(* Logix 5000 project; controller PLC_MCC1201_220AP1 vendor 1 type 14 code 164 rev 35.11; software revision 35.00 *)

TASK _18_STI (periodic, rate 10 ms, priority 10, watchdog 500 ms) : _18_STI
TASK Diagnostic (periodic, rate 500 ms, priority 15, watchdog 2000 ms) : Modules
TASK MainTask (periodic, rate 10 ms, priority 10, watchdog 500 ms) : MainProgram, CommandLogic

MODULES
   Local : vendor 1 type 14 code 164 (ICP 1, rev 35.11)
      PLC_MCC1300_TEST : vendor 1 type 14 code 166 (Ethernet 192.168.38.1, rev 35.1, $337b92f8$ RPI 20 ms)
      ETH_MCC1201 : 1756-EN2T (ICP 3, Ethernet 138.84.12.111, rev 11.1)
         Cullet_System : vendor 1 type 14 code 164 (Ethernet 138.84.12.122, rev 35.1, $37a2f589$ RPI 20 ms)
         ETH_MCC1300 : 1756-EN2T (Ethernet 138.84.12.118, rev 11.1, Output RPI 10 ms)
            PLC_MCC1300 : vendor 1 type 14 code 166 (ICP 0, rev 35.1)
      ETH_CULLET : 1756-EN2T (ICP 2, Ethernet 192.168.130.21, rev 11.1)
      A80AZ1 : PowerFlex 525-EENET (Ethernet 192.168.21.122, rev 7.1, Output RPI 20 ms)
      A81AZ1 : PowerFlex 525-EENET (Ethernet 192.168.21.123, rev 7.1, Output RPI 20 ms)
      PANEL_W2 : 1794-AENTR (Ethernet 192.168.24.62, rev 2.1, Output RPI 20 ms)
         R08_S01 : 1794-IB16 (Flex 1, rev 1.1)
         R08_S00 : 1794-IB16 (Flex 0, rev 1.1)
         R08_S02 : 1794-IB16 (Flex 2, rev 1.1)
         R08_S03 : vendor 1 type 7 code 35 (Flex 3, rev 1.1)
      CB_1CS : 1794-AENTR (Ethernet 192.168.24.51, rev 2.1, Output RPI 20 ms)
         R01_S00 : 1794-IB16 (Flex 0, rev 1.1)
         R01_S01 : vendor 1 type 7 code 35 (Flex 1, rev 1.1)
      CB_2CS : 1794-AENTR (Ethernet 192.168.24.52, rev 2.1, Output RPI 20 ms)
         R02_S00 : 1794-IB16 (Flex 0, rev 1.1)
         R02_S01 : vendor 1 type 7 code 35 (Flex 1, rev 1.1)
      CB_3CS : 1794-AENTR (Ethernet 192.168.24.53, rev 2.1, Output RPI 20 ms)
         R03_S00 : 1794-IB16 (Flex 0, rev 1.1)
         R03_S01 : vendor 1 type 7 code 35 (Flex 1, rev 1.1)
      CB_4CS : 1794-AENTR (Ethernet 192.168.24.54, rev 2.1, Output RPI 20 ms)
         R04_S00 : 1794-IB16 (Flex 0, rev 1.1)
         R04_S01 : vendor 1 type 7 code 35 (Flex 1, rev 1.1)
      CB_5CS : 1794-AENTR (Ethernet 192.168.24.55, rev 2.1, Output RPI 20 ms)
         R05_S00 : 1794-IB16 (Flex 0, rev 1.1)
         R05_S01 : vendor 1 type 7 code 35 (Flex 1, rev 1.1)
      MI_6CS : 1794-AENTR (Ethernet 192.168.24.56, rev 2.1, Output RPI 20 ms)
         R06_S00 : 1794-IB16 (Flex 0, rev 1.1)
         R06_S01 : vendor 1 type 7 code 35 (Flex 1, rev 1.1)
      PANEL_W3 : 1794-AENTR (Ethernet 192.168.24.63, rev 2.1, Output RPI 20 ms)
         R09_S01 : 1794-IB16 (Flex 1, rev 1.1)
         R09_S00 : 1794-IB16 (Flex 0, rev 1.1)
         R09_S03 : vendor 1 type 7 code 35 (Flex 3, rev 1.1)
         R09_S02 : 1794-IB16 (Flex 2, rev 1.1)
      A53AZ1 : vendor 1 type 45 code 15 (Ethernet 192.168.21.101, rev 2.3, AMotionDiagnostics RPI 1 ms)
      A54AZ1 : vendor 1 type 45 code 15 (Ethernet 192.168.21.102, rev 2.3, AMotionDiagnostics RPI 1 ms)
      A55AZ1 : vendor 1 type 45 code 15 (Ethernet 192.168.21.103, rev 2.3, AMotionDiagnostics RPI 1 ms)
      A61AZ1 : vendor 1 type 45 code 15 (Ethernet 192.168.21.105, rev 2.3, AMotionDiagnostics RPI 1 ms)
      A62AZ1 : vendor 1 type 45 code 15 (Ethernet 192.168.21.106, rev 2.3, AMotionDiagnostics RPI 1 ms)
      A63AZ1 : vendor 1 type 45 code 15 (Ethernet 192.168.21.107, rev 2.3, AMotionDiagnostics RPI 1 ms)
      A64AZ1 : vendor 1 type 45 code 15 (Ethernet 192.168.21.108, rev 2.3, AMotionDiagnostics RPI 1 ms)
      A65AZ1 : vendor 1 type 45 code 15 (Ethernet 192.168.21.109, rev 2.3, AMotionDiagnostics RPI 1 ms)
      A66AZ1 : vendor 1 type 45 code 15 (Ethernet 192.168.21.110, rev 2.3, AMotionDiagnostics RPI 1 ms)
      A67AZ1 : vendor 1 type 45 code 15 (Ethernet 192.168.21.111, rev 2.3, AMotionDiagnostics RPI 1 ms)
      A68AZ1 : vendor 1 type 45 code 15 (Ethernet 192.168.21.112, rev 2.3, AMotionDiagnostics RPI 1 ms)
      A69AZ1 : vendor 1 type 45 code 15 (Ethernet 192.168.21.113, rev 2.3, AMotionDiagnostics RPI 1 ms)
      A70AZ1 : vendor 1 type 45 code 15 (Ethernet 192.168.21.114, rev 2.3, AMotionDiagnostics RPI 1 ms)
      A71AZ1 : vendor 1 type 45 code 15 (Ethernet 192.168.21.115, rev 2.3, AMotionDiagnostics RPI 1 ms)
      A72AZ1 : vendor 1 type 45 code 15 (Ethernet 192.168.21.116, rev 2.3, AMotionDiagnostics RPI 1 ms)
      A73AZ1 : vendor 1 type 45 code 15 (Ethernet 192.168.21.117, rev 2.3, AMotionDiagnostics RPI 1 ms)
      A74AZ1 : vendor 1 type 45 code 15 (Ethernet 192.168.21.118, rev 2.3, AMotionDiagnostics RPI 1 ms)
      A77AZ1 : vendor 1 type 45 code 15 (Ethernet 192.168.21.121, rev 2.3, AMotionDiagnostics RPI 1 ms)
      A57AZ1 : vendor 1 type 45 code 15 (Ethernet 192.168.21.104, rev 2.3, AMotionDiagnostics RPI 1 ms)
      A75AZ1 : vendor 1 type 45 code 15 (Ethernet 192.168.21.119, rev 2.3, AMotionDiagnostics RPI 1 ms)
      A76AZ1 : vendor 1 type 45 code 15 (Ethernet 192.168.21.120, rev 2.3, AMotionDiagnostics RPI 1 ms)
      A155SW1 : vendor 1 type 12 code 246 (Ethernet 192.168.21.230, rev 12.1, Output RPI 1000 ms)
      A152AP1 : vendor 1 type 12 code 317 (Ethernet 192.168.21.11, rev 4.1)
         R00_S01 : 5069-IB16 (5069 1, rev 2.1, StandardDataDriven RPI 5 ms)
         R00_S02 : 5069-IB16 (5069 2, rev 2.1, StandardDataDriven RPI 5 ms)
         R00_S03 : 5069-IB16 (5069 3, rev 2.1, StandardDataDriven RPI 5 ms)
         R00_S04 : 5069-IB16 (5069 4, rev 2.1, StandardDataDriven RPI 5 ms)
         R00_S05 : 5069-IB16 (5069 5, rev 2.1, StandardDataDriven RPI 5 ms)
         R00_S06 : 5069-IB16 (5069 6, rev 2.1, StandardDataDriven RPI 5 ms)
         R00_S07 : 5069-IB16 (5069 7, rev 2.1, StandardDataDriven RPI 5 ms)
         R00_S08 : 5069-IB16 (5069 8, rev 2.1, StandardDataDriven RPI 5 ms)
         R00_S09 : 5069-IB16 (5069 9, rev 2.1, StandardDataDriven RPI 5 ms)
         R00_S10 : 5069-IB16 (5069 10, rev 2.1, StandardDataDriven RPI 5 ms)
         R00_S11 : 5069-IB16 (5069 11, rev 2.1, StandardDataDriven RPI 5 ms)
         R00_S12 : 5069-IB16 (5069 12, rev 2.1, StandardDataDriven RPI 5 ms)
         R00_S13 : 5069-OB16 (5069 13, rev 3.1, StandardDataDriven RPI 5 ms)
         R00_S14 : 5069-OB16 (5069 14, rev 3.1, StandardDataDriven RPI 5 ms)
         R00_S15 : 5069-OB16 (5069 15, rev 3.1, StandardDataDriven RPI 5 ms)
         R00_S16 : 5069-OB16 (5069 16, rev 3.1, StandardDataDriven RPI 5 ms)
         R00_S17 : 5069-OB16 (5069 17, rev 3.1, StandardDataDriven RPI 5 ms)
         R00_S18 : 5069-OB16 (5069 18, rev 3.1, StandardDataDriven RPI 5 ms)
END_MODULES

TYPE AOI_AccessArea_Alm :
STRUCT
   rgxS : AOI_AccessArea_StopFault;   // Stopping faults
   rgxF : AOI_AccessArea_Fault;   // Faults
   rgxW : AOI_AccessArea_Warning;   // Warnings
END_STRUCT
END_TYPE

TYPE AOI_AccessArea_Fault :   // Faults
STRUCT
   x0 : BOOL;   // Spare 0
   x1 : BOOL;   // Spare 1
   x2 : BOOL;   // Spare 2
   x3 : BOOL;   // Spare 3
   x4 : BOOL;   // Spare 4
   x5 : BOOL;   // Spare 5
   x6 : BOOL;   // Spare 6
   x7 : BOOL;   // Spare 7
   x8 : BOOL;   // Spare 8
   x9 : BOOL;   // Spare 9
   x10 : BOOL;   // Spare 10
   x11 : BOOL;   // Spare 11
   x12 : BOOL;   // Spare 12
   x13 : BOOL;   // Spare 13
   x14 : BOOL;   // Spare 14
   x15 : BOOL;   // Spare 15
   x16 : BOOL;   // Spare 16
   x17 : BOOL;   // Spare 17
   x18 : BOOL;   // Spare 18
   x19 : BOOL;   // Spare 19
   x20 : BOOL;   // Spare 20
   x21 : BOOL;   // Spare 21
   x22 : BOOL;   // Spare 22
   x23 : BOOL;   // Spare 23
   x24 : BOOL;   // Spare 24
   x25 : BOOL;   // Spare 25
   x26 : BOOL;   // Spare 26
   x27 : BOOL;   // Spare 27
   x28 : BOOL;   // Spare 28
   x29 : BOOL;   // Spare 29
   x30 : BOOL;   // Spare 30
   x31 : BOOL;   // Spare 31
END_STRUCT
END_TYPE

TYPE AOI_AccessArea_GP_STC :
STRUCT
   ST_xAccessRequest : BOOL;
   ST_xAccessAccepted : BOOL;
   ST_xAccessAnnulled : BOOL;
   ST_xAccessAcceptedAndButtonReleased : BOOL;
   ST_xDelayForceAccess : BOOL;
   ST_xSafetyOk : BOOL;
   OSR_xAccessRequest : BOOL;
   OSR_xAccessAcceptedAndButtonReleased : BOOL;
   OSR_xRemoveAccess : BOOL;
   OSR_xRemoveAccessNotAccepted : BOOL;
   OS_xAccessRequest : BOOL;
   OS_xSafetyOK : BOOL;
   tmON_ForceAccess : TIMER;
END_STRUCT
END_TYPE

TYPE AOI_AccessArea_HMR :
STRUCT
   dStatusAccessPoint : DINT;   // Status Door [1=OK; 7=Tripped] {x|x|x|x|O}
   dStatusAccessArea : DINT;   // Status Access Area [1=Area Ok; 2=Request ; 4=Acess Done; 8=Accepted] {x|x|x|x|O}
END_STRUCT
END_TYPE

TYPE AOI_AccessArea_StopFault :   // Stop Faults
STRUCT
   xSafety_Area_Intervened : BOOL;   // ##CONPONENT#.Safety Area Intervened
   x1 : BOOL;   // Spare 1
   x2 : BOOL;   // Spare 2
   x3 : BOOL;   // Spare 3
   x4 : BOOL;   // Spare 4
   x5 : BOOL;   // Spare 5
   x6 : BOOL;   // Spare 6
   x7 : BOOL;   // Spare 7
   x8 : BOOL;   // Spare 8
   x9 : BOOL;   // Spare 9
   x10 : BOOL;   // Spare 10
   x11 : BOOL;   // Spare 11
   x12 : BOOL;   // Spare 12
   x13 : BOOL;   // Spare 13
   x14 : BOOL;   // Spare 14
   x15 : BOOL;   // Spare 15
   x16 : BOOL;   // Spare 16
   x17 : BOOL;   // Spare 17
   x18 : BOOL;   // Spare 18
   x19 : BOOL;   // Spare 19
   x20 : BOOL;   // Spare 20
   x21 : BOOL;   // Spare 21
   x22 : BOOL;   // Spare 22
   x23 : BOOL;   // Spare 23
   x24 : BOOL;   // Spare 24
   x25 : BOOL;   // Spare 25
   x26 : BOOL;   // Spare 26
   x27 : BOOL;   // Spare 27
   x28 : BOOL;   // Spare 28
   x29 : BOOL;   // Spare 29
   x30 : BOOL;   // Spare 30
   x31 : BOOL;   // Spare 31
END_STRUCT
END_TYPE

TYPE AOI_AccessArea_STRUCT :
STRUCT
   tAlm : AOI_AccessArea_Alm;
   tHMR : AOI_AccessArea_HMR;
   tSTC : AOI_AccessArea_Logic;
END_STRUCT
END_TYPE

TYPE AOI_AccessArea_Warning :   // fault
STRUCT
   xRequestAccessAreaActive : BOOL;   // Spare 0
   xAccessAreaDone : BOOL;   // Spare 1
   x2 : BOOL;   // Spare 2
   x3 : BOOL;   // Spare 3
   x4 : BOOL;   // Spare 4
   x5 : BOOL;   // Spare 5
   x6 : BOOL;   // Spare 6
   x7 : BOOL;   // Spare 7
   x8 : BOOL;   // Spare 8
   x9 : BOOL;   // Spare 9
   x10 : BOOL;   // Spare 10
   x11 : BOOL;   // Spare 11
   x12 : BOOL;   // Spare 12
   x13 : BOOL;   // Spare 13
   x14 : BOOL;   // Spare 14
   x15 : BOOL;   // Spare 15
   x16 : BOOL;   // Spare 16
   x17 : BOOL;   // Spare 17
   x18 : BOOL;   // Spare 18
   x19 : BOOL;   // Spare 19
   x20 : BOOL;   // Spare 20
   x21 : BOOL;   // Spare 21
   x22 : BOOL;   // Spare 22
   x23 : BOOL;   // Spare 23
   x24 : BOOL;   // Spare 24
   x25 : BOOL;   // Spare 25
   x26 : BOOL;   // Spare 26
   x27 : BOOL;   // Spare 27
   x28 : BOOL;   // Spare 28
   x29 : BOOL;   // Spare 29
   x30 : BOOL;   // Spare 30
   x31 : BOOL;   // Spare 31
END_STRUCT
END_TYPE

TYPE DATA_TRACKING_RIBBON :
STRUCT
   dTotalAreaLength_cmm : DINT;   // Total area length [mm/100]
   dStepAdvancement_cmm : DINT;   // Step advancement [mm/100]
   dEncoderValueOnAdv_cmm : DINT;   // Encoder value on advancement [mm/100]
   dOperationInProgress : DINT;   // Task operation in progress
   rgtRibbons : DATA_TRACKING_RIBBON_DETAILS[200];   // Ribbon details
END_STRUCT
END_TYPE

TYPE DATA_TRACKING_RIBBON_DETAILS :
STRUCT
   rgxGlassBreak : DINT;   // Glass break info
   dGrossRibbonWidth_cmm : DINT;   // Gross ribbon width [mm/100]
   dNetRibbonWidth_cmm : DINT;   // Net ribbon width [mm/100]
   dGrossWander_cmm : DINT;   // Gross wander [mm/100]
   dNetWander_cmm : DINT;   // Net wander [mm/100]
END_STRUCT
END_TYPE

TYPE GP_AccessArea_STC :
STRUCT
   ST_xAccessRequest : BOOL;
   ST_xAccessAccepted : BOOL;
   ST_xAccessAnnulled : BOOL;
   ST_xAccessAcceptedAndButtonReleased : BOOL;
   ST_xConditionOkForAccess : BOOL;
   ST_xDelayForceAccess : BOOL;
   ST_xSafetyOkForCycle : BOOL;
   OSR_xAccessRequest : BOOL;
   OSR_xAccessAcceptedAndButtonReleased : BOOL;
   OSR_xRemoveAccess : BOOL;
   OSR_xRemoveAccessNotAccepted : BOOL;
   OS_xAccessRequest : BOOL;
   OS_xSafetyOK : BOOL;
   tmON_ForceAccess : TIMER;
END_STRUCT
END_TYPE

TYPE GP_NetworkDiag_v1 :
STRUCT
   sModuleName : STRING;   // Module name
   xConnected : BOOL;   // Module connected
   xFaulted : BOOL;   // Module faulted
   dEntryStatus : DINT;
   dFaultCode : DINT;
   dFaultInfo : DINT;
   dInstance : DINT;
END_STRUCT
END_TYPE

TYPE GP_OB_Initialize_STC :
STRUCT
   dElapsed_1h_ms : DINT; {access None}   // Decimal
   dElapsed_1min_ms : DINT; {access None}   // Decimal
   dElapsed_1s_ms : DINT; {access None}   // Decimal
   dElapsed_2min_ms : DINT; {access None}   // Decimal
   dElapsed_2s_ms : DINT; {access None}   // Decimal
   dElapsed_5s_ms : DINT; {access None}   // Decimal
   dElapsed_10min_ms : DINT; {access None}   // Decimal
   dElapsed_10s_ms : DINT; {access None}   // Decimal
   dElapsed_30min_ms : DINT; {access None}   // Decimal
   dElapsed_30s_ms : DINT; {access None}   // Decimal
   dElapsed_100ms_ms : DINT; {access None}   // Decimal
   dElapsed_200ms_ms : DINT; {access None}   // Decimal
   dElapsed_400ms_ms : DINT; {access None}   // Decimal
   dElapsed_500ms_ms : DINT; {access None}   // Decimal
   dElapsed_800ms_ms : DINT; {access None}   // Decimal
   dlLastExecValue_us : DINT; {access None}   // Decimal
   rReminder_ms : REAL; {access None}   // Float
   lwOldStartTime : DINT[2];   // Old start time execution
   lwStartTime : DINT[2];   // Start time execution
END_STRUCT
END_TYPE

TYPE MAC_BREAKER :
STRUCT
   ST_xOutputEnableBreaker : BOOL;   // Output enable breaker
   ST_xStoppingFaultsBreaker : BOOL;   // Cumulative of stopping faults breaker
   ST_xPhaseInProgress : BOOL;   // Phase in progress
   ST_xFaults : BOOL;   // Cumulative of faults
   ST_xStoppingFaults : BOOL;   // Cumulative of stopping faults
   ST_xWarnings : BOOL;   // Cumulative of warning
   ST_xBreakerRunningRequest : BOOL;   // Breaker running request
   OS_xStartBreakerInput : BOOL;   // OS.Start breaker input
   OS_xStopBreakerInput : BOOL;   // OS.Stop breaker input
   OS_xBreakerRunning : BOOL;   // OS.Breaker running
   OS_xCrusherStopAfterTimeout : BOOL;   // OS.Crusher stop after timeout
   OSR_xStartBreakerInput : BOOL;   // OSR.Start breaker input
   OSR_xStopBreakerInput : BOOL;   // OSR.Stop breaker input
   OSR_xBreakerRunning : BOOL;   // OSR.Breaker running
   OSR_xCrusherStopAfterTimeout : BOOL;   // OSR.Crusher stop after timeout
   INPUT_xFeedBackBreakerRotation : BOOL;   // Input.Feedback breaker rotation
   INPUT_xProtectionBreaker : BOOL;   // Input.Protection Breaker
   INPUT_xProtectionFan : BOOL;   // Input.Protection fan breaker
   INPUT_xFeedbackExclusionInductance : BOOL;   // Input.Feedback exclusion inductance
   INPUT_xStartBreaker : BOOL;   // Input.Start breaker
   INPUT_xStopBreaker : BOOL;   // Input.Stop breaker
   INPUT_xBreakerControlRotation : BOOL;   // Input.Breaker control rotation
   INPUT_xThermalProbe : BOOL;   // Input.Thermal probe
   INPUT_xLocalSafetySwitch : BOOL;   // Input.Local safety switch
   OUTPUT_xBreakerRun : BOOL;   // Output.Breaker run
   AUX_tmONCrusherStopDelayed : TIMER;   // Timer crusher stop delayed
   AUX_tmONFeedbackBreakerRot : TIMER;   // Timer feedback breaker rotation
   AUX_tmONBreakControlRotation : TIMER;   // Timer breaker control rotation
   AUX_tmONFeedbackBrakeBreakRot : TIMER;   // Timer feedback brake breaker rotation
   AUX_tmONFeedbackExclusionInduct : TIMER;   // Timer feedback inductance
END_STRUCT
END_TYPE

TYPE MAC_BREAKER_ALM :
STRUCT
   rgxStoppingFaults : DINT[2];   // Stopping faults
   rgxFaults : DINT[1];   // Faults
   rgxWarning : DINT[1];   // Warning
   rgdCodeAlarm : DINT[1];   // Code faults
END_STRUCT
END_TYPE

TYPE MAC_BREAKER_HMR :
STRUCT
   dBreakerStatus : DINT;   // Breaker status (1=Idle 3=Running 7=Anomaly) {x|x|x|x|O}
   xMan_BreakerRotateFdbk : BOOL;   // Manual breaker rotate fdbk {x|x|x|x|O}
END_STRUCT
END_TYPE

TYPE MAC_BREAKER_HMW :
STRUCT
   dTimeoutRunningCrusher_ms : DINT;   // Running crusher time [ms] {ms|s|0|3600|M}
   xMan_BreakerRotate : BOOL;   // Manual breaker rotate {x|x|x|x|O}
END_STRUCT
END_TYPE

TYPE MAC_CONVEYOR :
STRUCT
   ST_xOutputEnable : BOOL;   // Output enable
   ST_xPhaseInProgress : BOOL;   // Phase in progress
   ST_xFaults : BOOL;   // Cumulative of faults
   ST_xStoppingFaults : BOOL;   // Cumulative of stopping faults
   ST_xWarnings : BOOL;   // Cumulative of warning
   OUTPUT_xRun : BOOL;   // Output.Run
   OUTPUT_xDriveEnable : BOOL;   // Output.Drive enable
   OUTPUT_xDriveReset : BOOL;   // Output.Drive reset
   OUTPUT_xChangeSpeed : BOOL;   // Output.Drive change speed
   INPUT_xProtectionRot : BOOL;   // Input.Protection rotation
   INPUT_xProtectionFan : BOOL;   // Input.Protection fan rotation
   INPUT_xThermalProbe : BOOL;   // Input.Thermal probe
   INPUT_xDriveError : BOOL;   // Input.Drive error
   INPUT_xRotationFeedback : BOOL;   // Input.Rotation feedback
   INPUT_xDriveReady : BOOL;   // Input.Drive ready
   INPUT_xDriveInhibit : BOOL;   // Input.Drive inhibit
   INPUT_xLocalSafetySwitch : BOOL;   // Input.Local safety switch
   AUX_tmOFFRetainDriveEnable : TIMER;   // drive enable retain
   AUX_tmONRotfeedBackAlarm : TIMER;   // Rotation feedback alarm
   AUX_tmONDriveReadyAlarm : TIMER;   // Rotation feedback alarm
   OUTPUT_dSpeedReference_rpm : DINT;   // Output.Speed reference [rpm]
   AUX_rAcceleration_m_s2 : REAL;   // Acceleration [m/s2]
   AUX_rDeceleration_m_s2 : REAL;   // Deceleration [m/s2]
   AUX_dReqSpeed_mm_min : DINT;   // Request speed [mm/min]
   AUX_dRealSpeed_mm_min : DINT;   // Real speed [mm/min]
END_STRUCT
END_TYPE

TYPE MAC_CONVEYOR_ALM :
STRUCT
   rgxStoppingFaults : DINT[2];   // Stopping faults
   rgxFaults : DINT[1];   // Faults
   rgxWarning : DINT[1];   // Warning
   rgdCodeAlarm : DINT[1];   // Code faults
END_STRUCT
END_TYPE

TYPE MAC_CONVEYOR_HMR :
STRUCT
   xMan_JogForwardFdbk : BOOL;   // Manual jog forward fdbk {x|x|x|x|O}
   dStatus : DINT;   // Conveyor status (1=Idle 3=Running 7=Anomaly)
   dMode : DINT;   // Breaker Mode (1=Down; 2=Up; 4=Req Down; 8=Req Up) {X|X|X|X|O}
END_STRUCT
END_TYPE

TYPE MAC_CONVEYOR_HMW :
STRUCT
   xMan_JogForward : BOOL;   // Manual jog forward {x|x|x|x|O}
END_STRUCT
END_TYPE

TYPE MAC_CONVEYOR_IN_MOTION :
STRUCT
   DR_MAJ_M : MOTION_INSTRUCTION;   // Drive jog
   DR_MAS_M : MOTION_INSTRUCTION;   // Drive stop
END_STRUCT
END_TYPE

TYPE MAC_CONVEYOR_OUT_MOTION :
STRUCT
   DR_MSO_M : MOTION_INSTRUCTION;   // Drive ON
   DR_MSF_M : MOTION_INSTRUCTION;   // Drive OFF
   DR_MASR_M : MOTION_INSTRUCTION;   // Drive reset faults
   DR_MAJ_M : MOTION_INSTRUCTION;   // Drive jog
   DR_MCD_M : MOTION_INSTRUCTION;   // Drive change speed
   DR_MAS_M : MOTION_INSTRUCTION;   // Drive stop
END_STRUCT
END_TYPE

TYPE MAC_DROPCONV :
STRUCT
   ST_xOutputEnable : BOOL;   // Output enable
   ST_xPhaseInProgress : BOOL;   // Phase in progress
   ST_xFaults : BOOL;   // Cumulative of faults
   ST_xStoppingFaults : BOOL;   // Cumulative of stopping faults
   ST_xWarnings : BOOL;   // Cumulative of warning
   ST_xManualMode : BOOL;   // Manual mode
   OUTPUT_xRollerLifting : BOOL;   // Output.Roller lifting
   OUTPUT_xRiseDrop : BOOL;   // Output.Rise drop conveyor
   OUTPUT_xDescentDrop : BOOL;   // Output.Descent drop conveyor
   OUTPUT_xHLUpDownPushbutton : BOOL;   // Output.HL Up/Down pushbutton
   OUTPUT_xHLDoorOpenOpSide : BOOL;   // Output.HL Door open operator side
   OUTPUT_xHLDoorOpenFarSide : BOOL;   // Output.HL Door open far side
   INPUT_xProtection : BOOL;   // Input.Protection motor
   INPUT_xProtectionBrake : BOOL;   // Input.Protection brake
   INPUT_xFeedbackMovement : BOOL;   // Input.Movement feedback
   INPUT_xThermalProbe : BOOL;   // Input.Thermal probe
   INPUT_xUpPosition : BOOL;   // Input.Up position
   INPUT_xDownPosition : BOOL;   // Input.Down position
   INPUT_xFeedback : BOOL;   // Input.Movement feedback
   INPUT_xFeedbackBrake : BOOL;   // Input.Brake feedback
   INPUT_xTiltingSafetyBarDisinsered : BOOL;   // Input.Tilting Safety Bar Disinsered
   INPUT_xDoorOpenTiltingAreaOpSide : BOOL;   // Input.Door open tilting conveyor area operator side
   INPUT_xUpDownPushbuttonOpSide : BOOL;   // Input.Up/Down pushbutton operator side
   INPUT_xDoorOpenTiltingAreaFarSide : BOOL;   // Input.Door open tilting conveyor area far side
   INPUT_xUpDownPushbuttonFarSide : BOOL;   // Input.Up/Down pushbutton far side
   AUX_tmOFFEachCutAcceleration : TIMER;   // Acceleration time each cut
   AUX_tmOFFAcceleration : TIMER;   // Acceleration time
   AUX_tmONFeedbackMovAlarm : TIMER;   // Feedback movement alarm
   AUX_tmONFeedbackAlarm : TIMER;   // Feedback alarm
   AUX_tmONFeedbackBrakeAlarm : TIMER;   // Feedback brake alarm
   AUX_tmONMismatchSensorAlarm : TIMER;   // Mismatch sensor feedback alarm
   AUX_tmONUpSensorAlarm : TIMER;   // Up sensor feedback alarm
   AUX_tmONDownSensorAlarm : TIMER;   // Down sensor feedback alarm
   AUX_tmONForceUp : TIMER;   // Force up
   AUX_tmONEmCutTimeout : TIMER;   // Emergency Xcut timeout
   AUX_dDistanceToDescent_cmm : DINT;   // Distance to descent [mm/100]
   AUX_dDistanceToCheckGlass_cmm : DINT;   // Distance to check glass [mm/100]
   AUX_dConveyorLength_cmm : DINT;   // Conveyor length [mm/100]
   AUX_dAccelerationTime_ms : DINT;   // Acceleration time [ms]
   AUX_dAccelerationFactor : DINT;   // Acceleration factor
   AUX_dMaxSpeed_mm_min : DINT;   // Max speed [mm/min]
   AUX_dAccelerationSpeed_mm_min : DINT;   // Acceleration speed [mm/min]
   ST_xConditionOKforStopCycle : BOOL;   // Condition for stop cycle
   ST_xConveyorUpRequest : BOOL;   // Conveyor Up request
   ST_xConveyorDwRequest : BOOL;   // Conveyor Down request
   ST_xConveyorUp : BOOL;   // Conveyor Up
   ST_xUpFromPush : BOOL;   // Up from pushbutton
   ST_xUpFromScada : BOOL;   // Up from scada
   ST_xCutForQltPopup : BOOL;   // Cut arrived for qlt popup
   ST_xCutArrived : BOOL;   // Cut arrived
   ST_xXCutOffRequestAcceleration : BOOL;   // Emergency cut off - request acceleration
   ST_xEachCutAccelerationRequest : BOOL;   // Accelerate command for each cut request
   ST_xEachCutAcceleration : BOOL;   // Accelerate command for each cut
   ST_xAccelerateCommand : BOOL;   // Accelerate command
   ST_xEmCutArrived : BOOL;   // Emergency cut arrived (ready for descent)
   ST_xEmCutTimeout : BOOL;   // Emergency cut timeout
   OSR_xUpDownSBRequest : BOOL;   // OSR Up/Down pushbutton request
   OS_xUpDownSBRequest : BOOL;   // OS Up/Down pushbutton request
   OSR_xForceUpSBRequest : BOOL;   // OSR force up pushbutton request
   OS_xForceUpSBRequest : BOOL;   // OS force up pushbutton request
   OSR_xAccelerate : BOOL;   // OSR Accelerate
   OS_xAccelerate : BOOL;   // OS Accelerate
   OSR_xRise : BOOL;   // OSR Rise
   OS_xRise : BOOL;   // OS Rise
   OSR_xDescent : BOOL;   // OSR Descent
   OS_xDescent : BOOL;   // OS Descent
   OSR_xManCmdRise : BOOL;   // OSR Man Cmd Rise
   OS_xManCmdRise : BOOL;   // OS Man Cmd Rise
   OSR_xManCmdDescent : BOOL;   // OSR Man Cmd Descent
   OS_xManCmdDescent : BOOL;   // OS Man Cmd Descent
   OSR_xBreak : BOOL;   // OSR Glass break
   OSR_xCutForQltPopup : BOOL;   // OSR Cut for Qlt Popup
   OSR_xCutForQltPopupEnd : BOOL;   // OSR Cut for Qlt Popup end
END_STRUCT
END_TYPE

TYPE MAC_DROPCONV_ALM :
STRUCT
   rgxStoppingFaults : DINT[2];   // Stopping faults
   rgxFaults : DINT[1];   // Faults
   rgxWarning : DINT[1];   // Warning
   rgdCodeAlarm : DINT[1];   // Code faults
END_STRUCT
END_TYPE

TYPE MAC_DROPCONV_HMR :
STRUCT
   xMan_RiseFdbk : BOOL;   // Manual rise fdbk {x|x|x|x|O}
   xMan_DescentFdbk : BOOL;   // Manual descent fdbk {x|x|x|x|O}
   xUpPosition : BOOL;   // Up position {x|x|x|x|O}
   xDownPosition : BOOL;   // Down position {x|x|x|x|O}
   xEnabledBreakingDetection : BOOL;   // Enabled automatic descent for glass break {x|x|x|x|O}
   xDoorOpenedOperatorSide : BOOL;   // Door opened operator side {x|x|x|x|O}
   xDoorOpenedFarSide : BOOL;   // Door opened far side {x|x|x|x|O}
   dMode : DINT;   // Drop mode (1=Down 2=Up 4=Req Down 8=Req up)
   dStatus : DINT;   // Drop conveyor status (1=Idle 3=Moving 7=Anomaly)
   dDistanceFromSnaproll_cmm : DINT;   // Distance from snaproll [mm/100] {mm/100|mm|x|x|O}
END_STRUCT
END_TYPE

TYPE MAC_DROPCONV_HMW :
STRUCT
   xMan_Rise : BOOL;   // Manual rise {x|x|x|x|O}
   xMan_Descent : BOOL;   // Manual descent {x|x|x|x|O}
   dDistanceFromSnaproll_cmm : DINT;   // Distance from snaproll [mm/100] {mm/100|mm|0|65000|M}
   xUpdateDistanceFromSnaproll : BOOL;   // Update distance from snaproll {x|x|x|x|M}
   xEnableBreakingDetection : BOOL;   // Enable automatic descent for glass break {x|x|x|x|O}
   xDisableBreakingDetection : BOOL;   // Disable automatic descent for glass break {x|x|x|x|O}
   xRequestUp : BOOL;   // Request tilting up {x|x|x|x|M}
   xRequestDown : BOOL;   // Request tilting down {x|x|x|x|M}
   xForceUp : BOOL;   // Force tilting up {x|x|x|x|M}
   xForceDown : BOOL;   // Force tilting down {x|x|x|x|M}
END_STRUCT
END_TYPE

TYPE MAC_EMERGENCYXCUT :
STRUCT
   ST_xOutputEnable : BOOL;   // Output enable
   ST_xAccessAreaRequestOpSide : BOOL;   // Access area request operator side
   ST_xAccessAreaRequestFarSide : BOOL;   // Access area request far side
   ST_xConditionOKAccessArea : BOOL;   // Condition ok for area access
   ST_xSelectorAutomaticMode : BOOL;   // Selector automatic mode
   ST_xSelectorManualMode : BOOL;   // Selector manual mode
   ST_xSemiautoModeSelection : BOOL;   // Semiauto mode selection
   ST_xAutomaticModeSelection : BOOL;   // Automatic mode selection
   ST_xManualModeSelection : BOOL;   // Manual mode selection
   ST_xManualModeAccepted : BOOL;   // Manual mode Accepted
   ST_xManualModeRequest : BOOL;   // Manual mode request
   ST_xSemiautoModeRequest : BOOL;   // Semiauto mode request
   ST_xSemiautoModeAccepted : BOOL;   // Semiauto mode accepted
   ST_xAutomaticModeAccepted : BOOL;   // Automatic mode accepted
   ST_xSemiautoMode : BOOL;   // Semiautomatic mode
   ST_xStopCycleRequest : BOOL;   // Stop cycle request continuous mode
   ST_xStartCycleRequest : BOOL;   // Start cycle request continuous mode
   ST_xStopCycleAccepted : BOOL;   // Stop cycle accepted
   ST_xCycleON : BOOL;   // Cycle ON continuous mode
   ST_xCondOKContinuousEmergencyCutting : BOOL;   // Condition OK Continuous mode cutting
   ST_xContinuousEmergencyCutting : BOOL;   // Continuous mode cutting
   ST_xSingleCuttingRequested : BOOL;   // Single cutting requested
   ST_xHeadDescent : BOOL;   // Head descent
   ST_xDistanceBetweenCutOK : BOOL;   // Distance between cut OK
   ST_xConditionOKLowerHead : BOOL;   // Condition OK to lower head
   ST_xConditionOKStopCycle : BOOL;   // Condition OK for stop cycle
   ST_xConditionOKCycleON : BOOL;   // Condition OK for cycle ON
   ST_xConditionOKSemiautoMode : BOOL;   // Condition OK for semiautomatic mode
   ST_xConditionOKManualMode : BOOL;   // Condition OK for manual mode
   ST_xMachineHomed : BOOL;   // Machine homed
   ST_xHeadDescentOneTime : BOOL;   // Head descent at least one time after rising
   ST_xCutDone : BOOL;   // Cut done
   ST_xBackwardPositionReached : BOOL;   // Backward position reached
   ST_xForwardPositionReached : BOOL;   // Forward position reached
   ST_xBreakerCutRequest : BOOL;   // Cut request coming from breaker
   ST_xPhaseInProgress : BOOL;   // Phase in progress
   ST_xFaults : BOOL;   // Cumulative of faults
   ST_xStoppingFaults : BOOL;   // Cumulative of stopping faults
   ST_xWarnings : BOOL;   // Cumulative of warning
   PH_xMoveForward : BOOL;   // Move fw
   PH_xEndMoveForward : BOOL;   // End Move fw
   PH_xMoveBackward : BOOL;   // Move bw
   PH_xEndMoveBackward : BOOL;   // End Move bw
   PH_xHoming : BOOL;   // Execute homing
   PH_xEndHoming : BOOL;   // End Execute homing
   OUTPUT_xJogFW : BOOL;   // Output.Run fw
   OUTPUT_xJogBW : BOOL;   // Output.Run bw
   OUTPUT_xHoming : BOOL;   // Output.Execute homing
   OUTPUT_xPositioning : BOOL;   // Output.Execute positioning
   OUTPUT_xDriveEnable : BOOL;   // Output.Drive enable
   OUTPUT_xMachineReady : BOOL;   // Output.HL Machine ready (Green)
   OUTPUT_xMachineToMaintenance : BOOL;   // Output.HL Machine to maintenance (Yellow)
   OUTPUT_xMachineOutOfOrder : BOOL;   // Output.HL Machine out of order (Red)
   OUTPUT_xAreaAccessRequestOpSide : BOOL;   // Output.HL Area access request operator side
   OUTPUT_xAreaAccessRequestFarSide : BOOL;   // Output.HL Area access request far side
   OUTPUT_xAreaSafetyOn : BOOL;   // Output.HL Area safety on
   OUTPUT_xUnlockDoorOpSide : BOOL;   // Output.Unlock safety door operator side
   OUTPUT_xUnlockDoorFarSide : BOOL;   // Output.Unlock safety door far side
   OUTPUT_xAutomatic : BOOL;   // Output.HL Automatic
   OUTPUT_xStartCut : BOOL;   // Output.HL Start cutting
   OUTPUT_xStopCut : BOOL;   // Output.HL Stop cutting
   OUTPUT_xCuttingHeadDescent : BOOL;   // Output.YV cutting head descent
   OUTPUT_xLubrication : BOOL;   // Output.YV lubrication
   OUTPUT_xAirActivation : BOOL;   // Output.YV air activation
   OUTPUT_xCarriageOverstroke : BOOL;   // Output.HL Carriage overstroke initial reset
   INPUT_xProtectionTraslation : BOOL;   // Input.Protection traslation
   INPUT_xProtectionFan : BOOL;   // Input.Protection fan rotation
   INPUT_xBreakingResTProbe : BOOL;   // Input.Breaking resistance thermal probe
   INPUT_xThermalProbe : BOOL;   // Input.Thermal probe
   INPUT_xDriveError : BOOL;   // Input.Drive error
   INPUT_xTraslationFeedback : BOOL;   // Input.Traslation feedback
   INPUT_xDriveReady : BOOL;   // Input.Drive ready
   INPUT_xAreaSafety : BOOL;   // Input.Area safety
   INPUT_xAccessAreaRequestOpSide : BOOL;   // Input.Area access request operator side
   INPUT_xResetAreaSafetiesOpSide : BOOL;   // Input.Reset area safeties operator side
   INPUT_xAccessAreaRequestFarSide : BOOL;   // Input.Area access request far side
   INPUT_xResetAreaSafetiesFarSide : BOOL;   // Input.Reset area safeties far side
   INPUT_xOverstrokeFW : BOOL;   // Input.Overstroke FW
   INPUT_xOverstrokeBW : BOOL;   // Input.Overstroke BW
   INPUT_xManual : BOOL;   // Input.Manual
   INPUT_xAutomatic : BOOL;   // Input.Automatic
   INPUT_xCutInterruption : BOOL;   // Input.Cutting interruption
   INPUT_xStartCut : BOOL;   // Input.Start cutting
   INPUT_xStopCut : BOOL;   // Input.Stop cutting
   INPUT_xAlarmOff : BOOL;   // Input.Alarm OFF
   INPUT_xLocalSafetySwitch : BOOL;   // Input.Local safety switch
   INPUT_xHomePosition : BOOL;   // Input.Home Position
   INPUT_xCompressedAirPresence : BOOL;   // Input.Compressed air presence
   INPUT_xLubricationTest : BOOL;   // Input.Lubrication test
   INPUT_xCuttingHeadTest : BOOL;   // Input.Cutting head test
   INPUT_xCuttingHeadHigh : BOOL;   // Input.Cutting head high
   INPUT_xCuttingSafety : BOOL;   // Input.Cutting safety
   INPUT_xOpeningDoorLocalizationOpSide : BOOL;   // Input.Opening door localization operator side
   INPUT_xOpeningDoorLocalizationFarSide : BOOL;   // Input.Opening door localization far side
   AUX_xHMIReqAutoPosition : BOOL;   // Request tilting auto position
   AUX_xHMIReqForceDown : BOOL;   // Request tilting force down
   AUX_dDistanceFTCHead : DINT;   // Distance from photocell to cutting head
   AUX_dBridgeAngle : DINT;   // Bridge angle [°/10000]
   AUX_dManualSpeed_mm_min : DINT;   // Manual mode speed [mm/min]
   AUX_dRiseReactionTime_ms : DINT;   // Rise reaction time [ms]
   AUX_dDescentReactionTime_ms : DINT;   // Descent reaction time [ms]
   AUX_dBackwardFastSpeed_mm_min : DINT;   // Return speed fast [mm/min]
   AUX_dBackwardSlowSpeed_mm_min : DINT;   // Return speed slow [mm/min]
   AUX_dCarriageInitialPosition_cmm : DINT;   // Carriage backward position [mm/100]
   AUX_dCarriageFinalPosition_cmm : DINT;   // Carriage forward position [mm/100]
   AUX_dMinimumStripeLength : DINT;   // Minimum stripe length [mm/100]
   AUX_dMaximumStripeLength : DINT;   // Maximum stripe length [mm/100]
   AUX_dTankElementCounter : DINT;   // Number of element on cut tank
   AUX_rgdCutTank : DINT[20];   // Tank encoder value on last cut
   AUX_dLastCutValue : DINT;   // Last cut encoder value
   AUX_dLastCutValueStored : DINT;   // Last cut encoder value
   AUX_dCutSpeed_mm_min : DINT;   // Cut speed [mm/min]
   AUX_dForwardTimeoutTime_ms : DINT;   // Timeout time forward phase [ms]
   AUX_dReturnSpeed_mm_min : DINT;   // Return speed [mm/min]
   AUX_dReqSpeed_mm_min : DINT;   // Speed request [mm/min]
   AUX_dStartControlPhotocellPos_dmm : DINT;   // Start control photocell position [mm/10]
   AUX_dTimeFTCToHead_ms : DINT;   // Time from photocel to head [ms]
   AUX_dTimeDelayToDescent_ms : DINT;   // Time delay to descent [ms]
   AUX_dTimeAdvanceToRise_ms : DINT;   // Time advance rise [ms]
   AUX_dTimeDelayToLubrication_ms : DINT;   // Time delay to lubricate ms]
   AUX_dTimeAdvanceToLubrication_ms : DINT;   // Time advance to lubricate [ms]
   OSR_xConditionNotOKToCut : BOOL;   // OSR condition not OK to cut
   OSR_xConditionNotAllowedLower : BOOL;   // OSR condition not allowed to lower head
   OSR_xSaveEncoderValue : BOOL;   // OSR save encoder value
   OSR_xRequestAccessAreaOpSide : BOOL;   // OSR access area request operator side
   OSR_xRequestAccessAreaFarSide : BOOL;   // OSR access area request far side
   OSR_xAreaSafetyOK : BOOL;   // OSR area safety ok
   OSR_xAreaSafety : BOOL;   // OSR area safety
   OSR_xStartCycle : BOOL;   // OSR start cycle
   OSR_xDriveHomed : BOOL;   // OSR drive homed